(* Logix 5000 project; controller MV vendor 1 type 14 code 217 rev 31.11; software revision 31.00; part 40 of 53 *)
(* tags used below, declared in another part *)
   active : BOOL;
   MV_B100 : INT[255];   // AT FLAGS
   MV_N101 : INT[255];   // AT INT Fermentation control integer workspace
   MV_N110 : INT[255];   // MV DATA 0 CURRENT FV DATA
   MV_N12 : INT[255];   // SYS_PARMS System Parameter Fil e
   MV_N14 : INT[255];   // ME>PLC Inter PLC comms traf fic outbound
   MV_N7 : INT[255];   // INTEGER
   MV_SFile : INT[255];   // SLC Equivalent System File, So Original Code Can Remain
   MV_T102 : TIMER[10];
   MV_T4 : TIMER[20];
   MV_TENTH_HOUR_OUTPUT_BIT : BOOL;
   temp : INT;
(* MV_Common, continued *)

ROUTINE MV_FV_ELAPSED_102   (* ladder *)
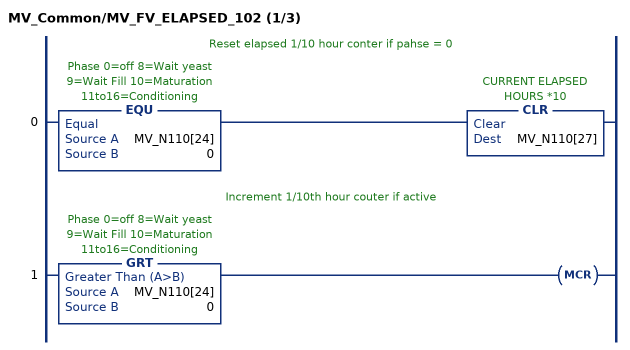
   // Reset elapsed 1/10 hour conter if pahse = 0
   0: EQU(MV_N110[24],0)CLR(MV_N110[27]);
   // Increment 1/10th hour couter if active
   1: GRT(MV_N110[24],0)MCR();
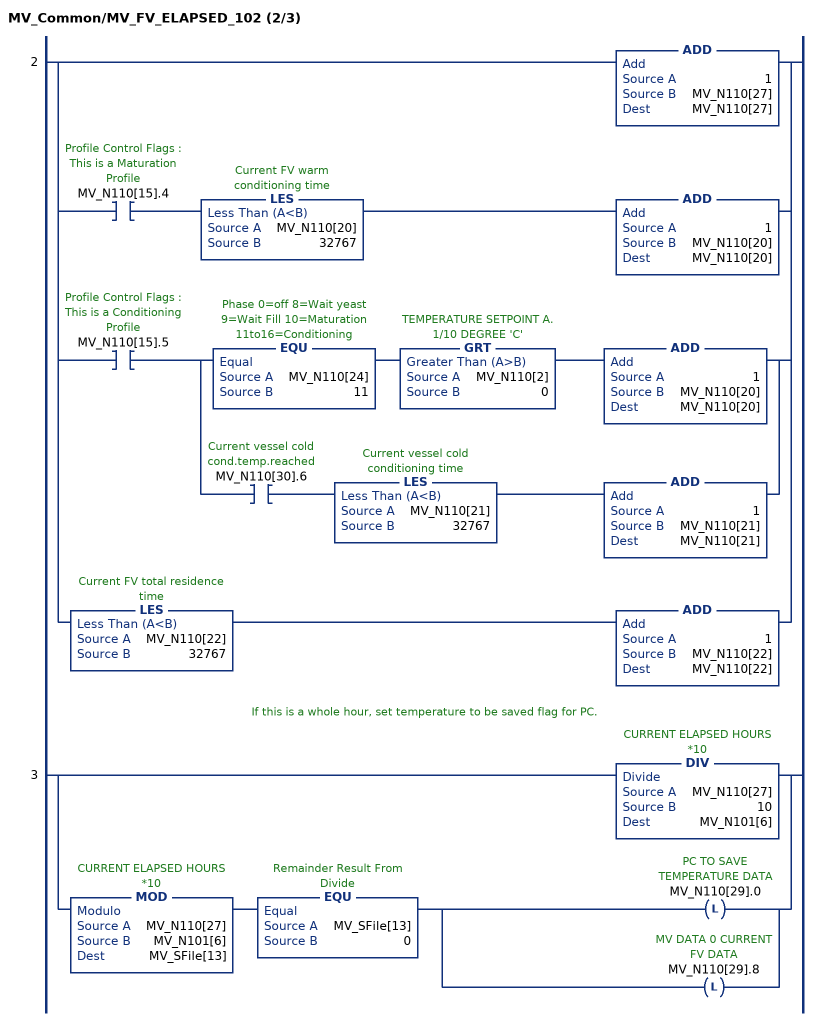
   2: [ADD(1,MV_N110[27],MV_N110[27]) ,XIC(MV_N110[15].4) LES(MV_N110[20],32767) ADD(1,MV_N110[20],MV_N110[20]) ,XIC(MV_N110[15].5) [EQU(MV_N110[24],11) GRT(MV_N110[2],0) ADD(1,MV_N110[20],MV_N110[20]) ,XIC(MV_N110[30].6) LES(MV_N110[21],32767) ADD(1,MV_N110[21],MV_N110[21]) ] ,LES(MV_N110[22],32767) ADD(1,MV_N110[22],MV_N110[22]) ];
   // If this is a whole hour, set temperature to be saved flag for PC.
   3: [DIV(MV_N110[27],10,MV_N101[6]) ,MOD(MV_N110[27],MV_N101[6],MV_SFile[13]) EQU(MV_SFile[13],0) [OTL(MV_N110[29].0) ,OTL(MV_N110[29].8) ] ];
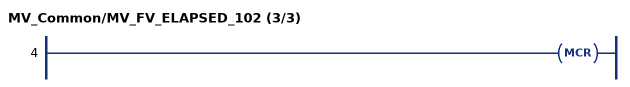
   4: MCR();
END_ROUTINE

ROUTINE MV_FV_MCP_100   (* ladder *)
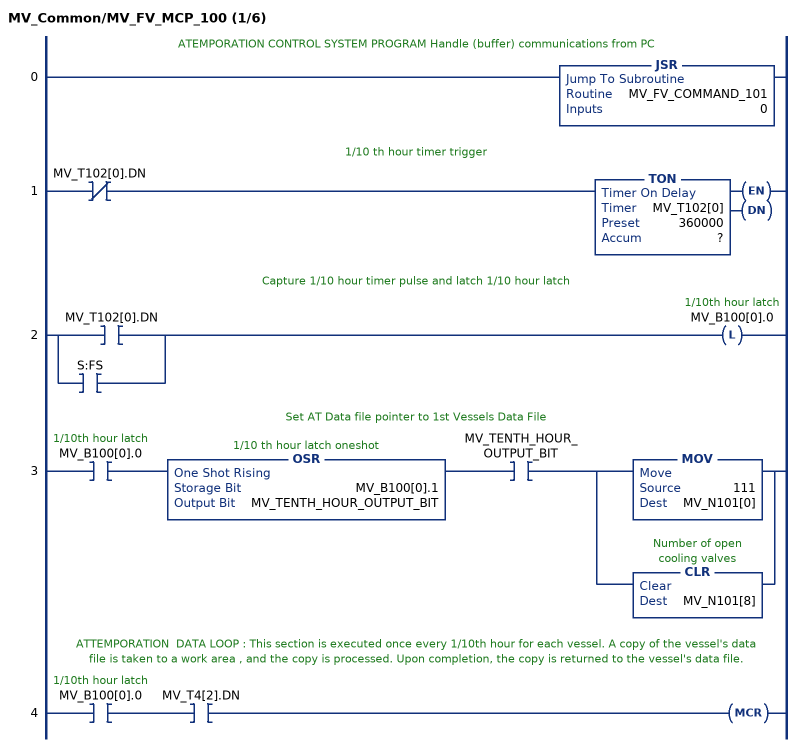
   // ATEMPORATION CONTROL SYSTEM PROGRAM Handle (buffer) communications from PC
   0: JSR(MV_FV_COMMAND_101,0);
   // 1/10 th hour timer trigger
   1: XIO(MV_T102[0].DN)TON(MV_T102[0],?,?);
   // Capture 1/10 hour timer pulse and latch 1/10 hour latch
   2: [XIC(MV_T102[0].DN) ,XIC(S:FS) ]OTL(MV_B100[0].0);
   // Set AT Data file pointer to 1st Vessels Data File
   3: XIC(MV_B100[0].0)OSR(MV_B100[0].1,MV_TENTH_HOUR_OUTPUT_BIT)XIC(MV_TENTH_HOUR_OUTPUT_BIT)[MOV(111,MV_N101[0]) ,CLR(MV_N101[8]) ];
   // ATTEMPORATION  DATA LOOP : This section is executed once every 1/10th hour for each vessel. A copy of the vessel's data file is taken to a work area , and the copy is processed. Upon completion, the copy is returned to the vessel's data file.
   4: XIC(MV_B100[0].0)XIC(MV_T4[2].DN)MCR();
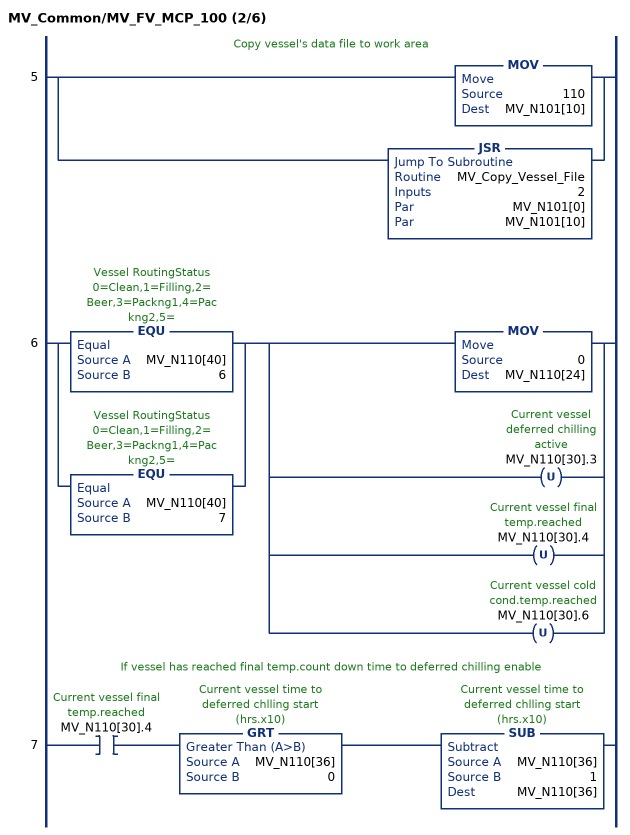
   // Copy vessel's data file to work area
   5: [MOV(110,MV_N101[10]) ,JSR(MV_Copy_Vessel_File,2,MV_N101[0],MV_N101[10]) ];
   6: [EQU(MV_N110[40],6) ,EQU(MV_N110[40],7) ][MOV(0,MV_N110[24]) ,OTU(MV_N110[30].3) ,OTU(MV_N110[30].4) ,OTU(MV_N110[30].6) ];
   // If vessel has reached final temp.count down time to deferred chilling enable
   7: XIC(MV_N110[30].4)GRT(MV_N110[36],0)SUB(MV_N110[36],1,MV_N110[36]);
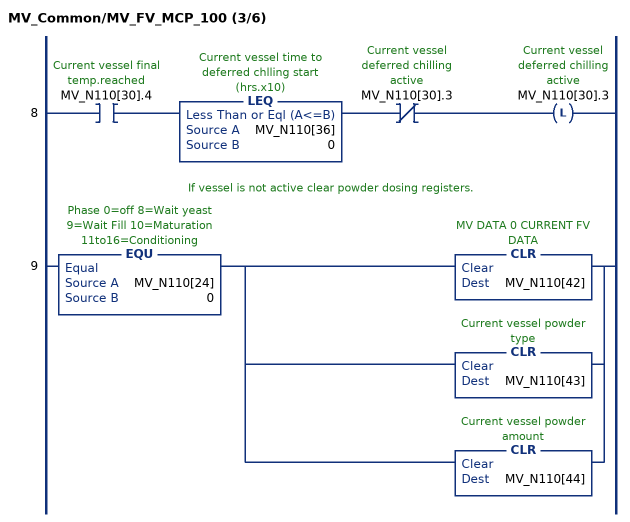
   8: XIC(MV_N110[30].4)LEQ(MV_N110[36],0)XIO(MV_N110[30].3)OTL(MV_N110[30].3);
   // If vessel is not active clear powder dosing registers.
   9: EQU(MV_N110[24],0)[CLR(MV_N110[42]) ,CLR(MV_N110[43]) ,CLR(MV_N110[44]) ];
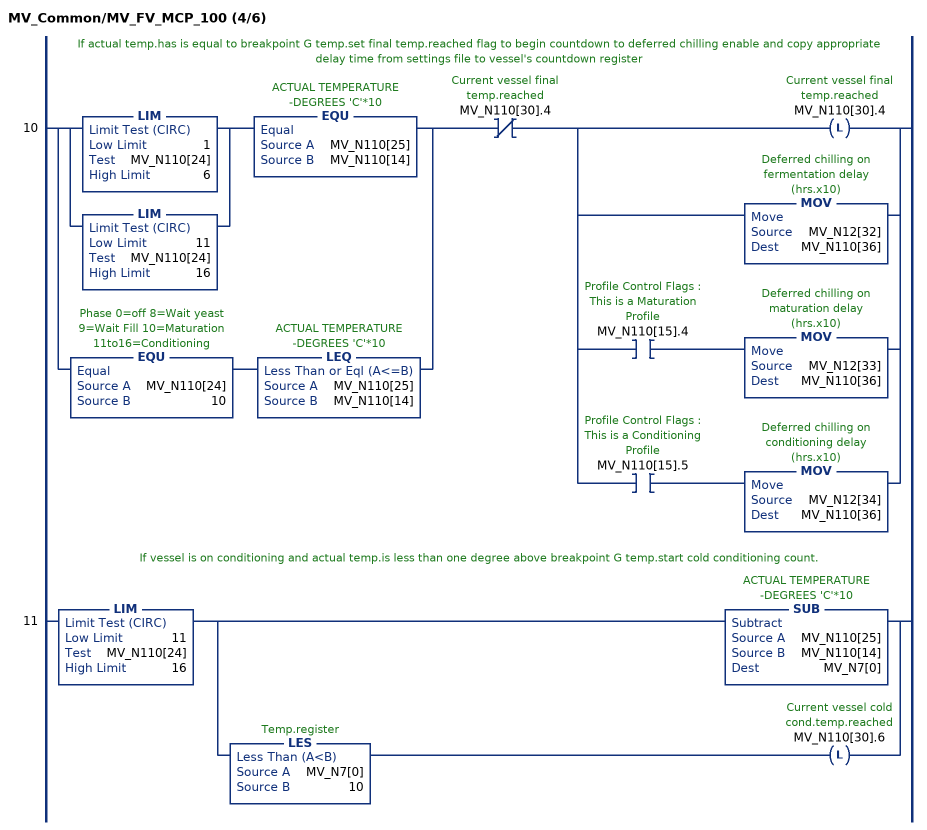
   // If actual temp.has is equal to breakpoint G temp.set final temp.reached flag to begin countdown to deferred chilling enable and copy appropriate delay time from settings file to vessel's countdown register
   10: [[LIM(1,MV_N110[24],6) ,LIM(11,MV_N110[24],16) ] EQU(MV_N110[25],MV_N110[14]) ,EQU(MV_N110[24],10) LEQ(MV_N110[25],MV_N110[14]) ]XIO(MV_N110[30].4)[OTL(MV_N110[30].4) ,MOV(MV_N12[32],MV_N110[36]) ,XIC(MV_N110[15].4) MOV(MV_N12[33],MV_N110[36]) ,XIC(MV_N110[15].5) MOV(MV_N12[34],MV_N110[36]) ];
   // If vessel is on conditioning and actual temp.is less than one degree above breakpoint G temp.start cold conditioning count.
   11: LIM(11,MV_N110[24],16)[SUB(MV_N110[25],MV_N110[14],MV_N7[0]) ,LES(MV_N7[0],10) OTL(MV_N110[30].6) ];
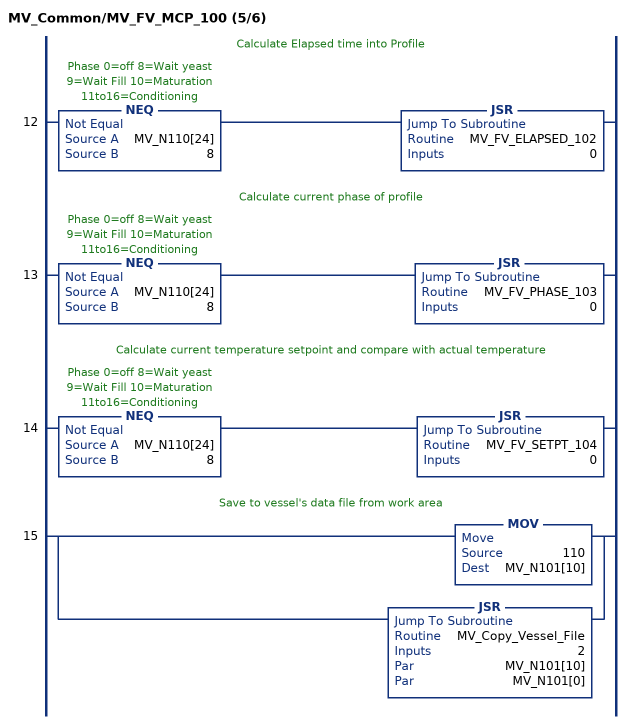
   // Calculate Elapsed time into Profile
   12: NEQ(MV_N110[24],8)JSR(MV_FV_ELAPSED_102,0);
   // Calculate current phase of profile
   13: NEQ(MV_N110[24],8)JSR(MV_FV_PHASE_103,0);
   // Calculate current temperature setpoint and compare with actual temperature
   14: NEQ(MV_N110[24],8)JSR(MV_FV_SETPT_104,0);
   // Save to vessel's data file from work area
   15: [MOV(110,MV_N101[10]) ,JSR(MV_Copy_Vessel_File,2,MV_N101[10],MV_N101[0]) ];
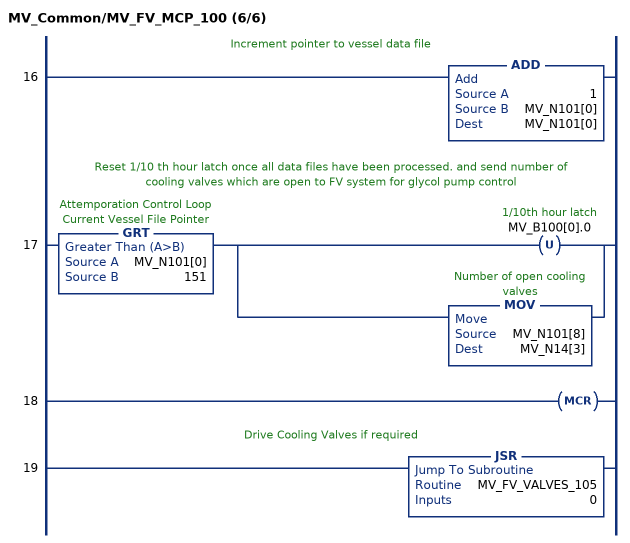
   // Increment pointer to vessel data file
   16: ADD(1,MV_N101[0],MV_N101[0]);
   // Reset 1/10 th hour latch once all data files have been processed. and send number of cooling valves which are open to FV system for glycol pump control
   17: GRT(MV_N101[0],151)[OTU(MV_B100[0].0) ,MOV(MV_N101[8],MV_N14[3]) ];
   18: MCR();
   // Drive Cooling Valves if required
   19: JSR(MV_FV_VALVES_105,0);
END_ROUTINE

ROUTINE MV_FV_PHASE_103   (* ladder *)
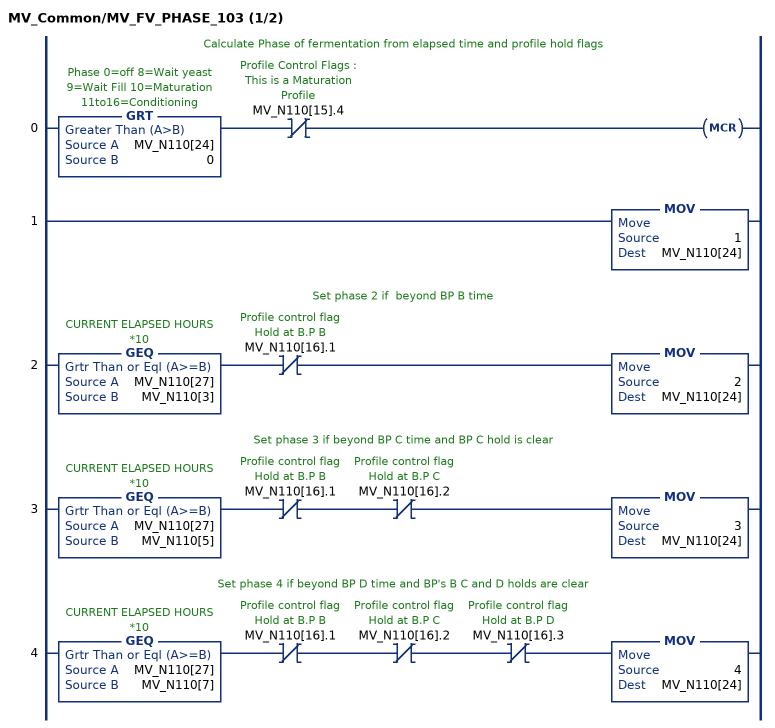
   // Calculate Phase of fermentation from elapsed time and profile hold flags
   0: GRT(MV_N110[24],0)XIO(MV_N110[15].4)MCR();
   1: MOV(1,MV_N110[24]);
   // Set phase 2 if  beyond BP B time
   2: GEQ(MV_N110[27],MV_N110[3])XIO(MV_N110[16].1)MOV(2,MV_N110[24]);
   // Set phase 3 if beyond BP C time and BP C hold is clear
   3: GEQ(MV_N110[27],MV_N110[5])XIO(MV_N110[16].1)XIO(MV_N110[16].2)MOV(3,MV_N110[24]);
   // Set phase 4 if beyond BP D time and BP's B C and D holds are clear
   4: GEQ(MV_N110[27],MV_N110[7])XIO(MV_N110[16].1)XIO(MV_N110[16].2)XIO(MV_N110[16].3)MOV(4,MV_N110[24]);
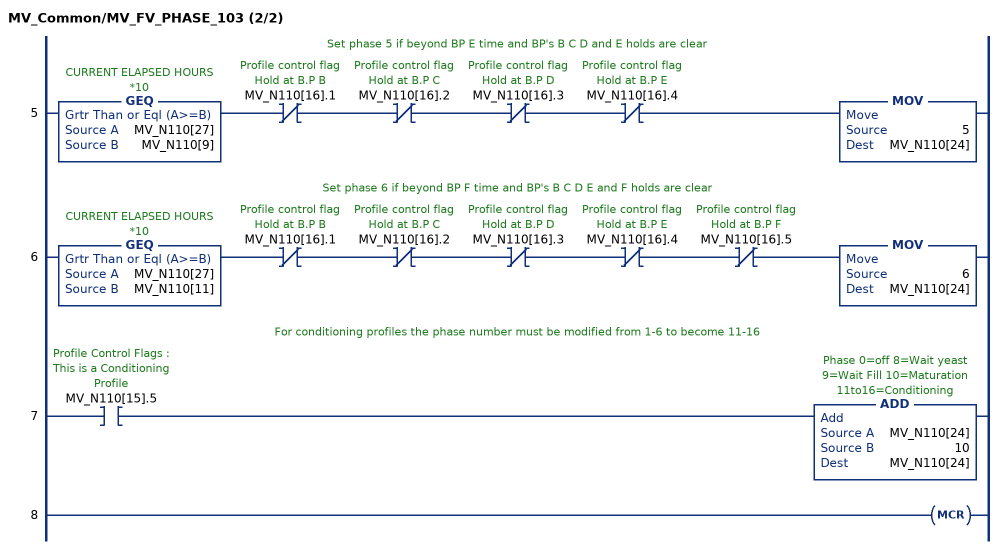
   // Set phase 5 if beyond BP E time and BP's B C D and E holds are clear
   5: GEQ(MV_N110[27],MV_N110[9])XIO(MV_N110[16].1)XIO(MV_N110[16].2)XIO(MV_N110[16].3)XIO(MV_N110[16].4)MOV(5,MV_N110[24]);
   // Set phase 6 if beyond BP F time and BP's B C D E and F holds are clear
   6: GEQ(MV_N110[27],MV_N110[11])XIO(MV_N110[16].1)XIO(MV_N110[16].2)XIO(MV_N110[16].3)XIO(MV_N110[16].4)XIO(MV_N110[16].5)MOV(6,MV_N110[24]);
   // For conditioning profiles the phase number must be modified from 1-6 to become 11-16
   7: XIC(MV_N110[15].5)ADD(MV_N110[24],10,MV_N110[24]);
   8: MCR();
END_ROUTINE

ROUTINE MV_FV_SETPT_104   (* ladder *)
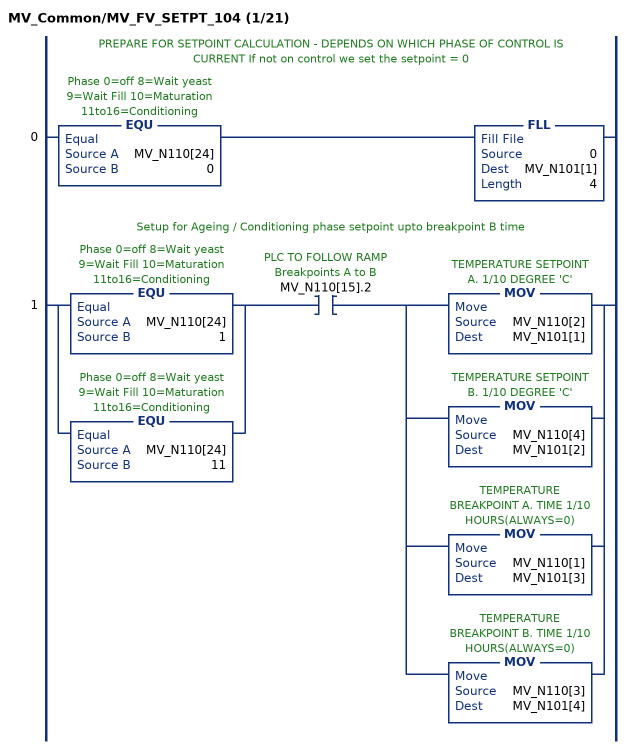
   // PREPARE FOR SETPOINT CALCULATION - DEPENDS ON WHICH PHASE OF CONTROL IS CURRENT If not on control we set the setpoint = 0
   0: EQU(MV_N110[24],0)FLL(0,MV_N101[1],4);
   // Setup for Ageing / Conditioning phase setpoint upto breakpoint B time
   1: [EQU(MV_N110[24],1) ,EQU(MV_N110[24],11) ]XIC(MV_N110[15].2)[MOV(MV_N110[2],MV_N101[1]) ,MOV(MV_N110[4],MV_N101[2]) ,MOV(MV_N110[1],MV_N101[3]) ,MOV(MV_N110[3],MV_N101[4]) ];
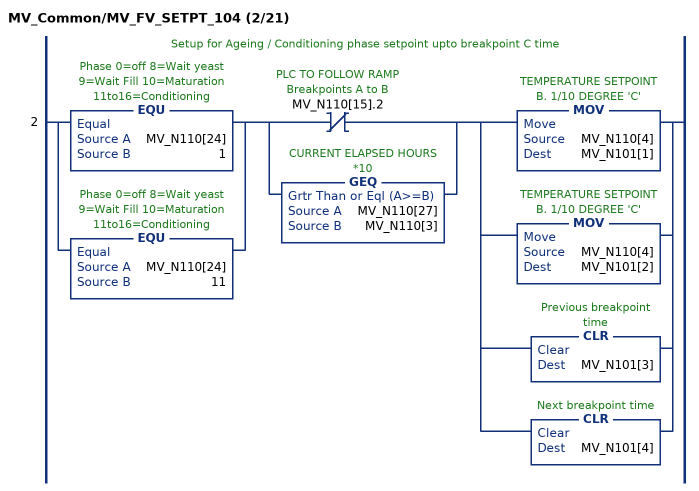
   // Setup for Ageing / Conditioning phase setpoint upto breakpoint C time
   2: [EQU(MV_N110[24],1) ,EQU(MV_N110[24],11) ][XIO(MV_N110[15].2) ,GEQ(MV_N110[27],MV_N110[3]) ][MOV(MV_N110[4],MV_N101[1]) ,MOV(MV_N110[4],MV_N101[2]) ,CLR(MV_N101[3]) ,CLR(MV_N101[4]) ];
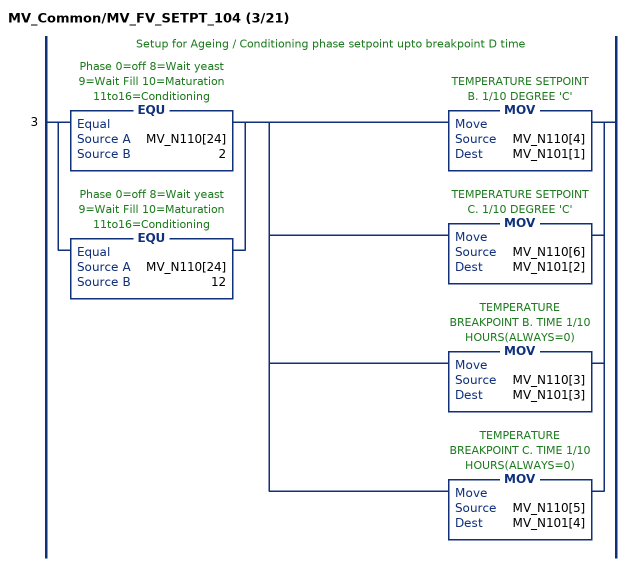
   // Setup for Ageing / Conditioning phase setpoint upto breakpoint D time
   3: [EQU(MV_N110[24],2) ,EQU(MV_N110[24],12) ][MOV(MV_N110[4],MV_N101[1]) ,MOV(MV_N110[6],MV_N101[2]) ,MOV(MV_N110[3],MV_N101[3]) ,MOV(MV_N110[5],MV_N101[4]) ];
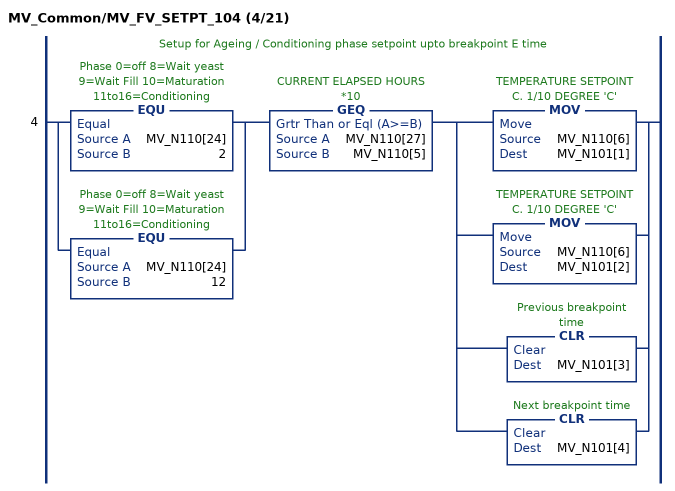
   // Setup for Ageing / Conditioning phase setpoint upto breakpoint E time
   4: [EQU(MV_N110[24],2) ,EQU(MV_N110[24],12) ]GEQ(MV_N110[27],MV_N110[5])[MOV(MV_N110[6],MV_N101[1]) ,MOV(MV_N110[6],MV_N101[2]) ,CLR(MV_N101[3]) ,CLR(MV_N101[4]) ];
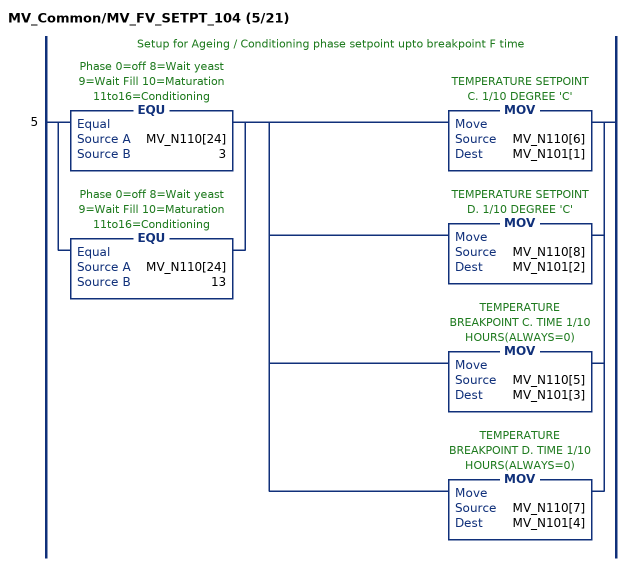
   // Setup for Ageing / Conditioning phase setpoint upto breakpoint F time
   5: [EQU(MV_N110[24],3) ,EQU(MV_N110[24],13) ][MOV(MV_N110[6],MV_N101[1]) ,MOV(MV_N110[8],MV_N101[2]) ,MOV(MV_N110[5],MV_N101[3]) ,MOV(MV_N110[7],MV_N101[4]) ];
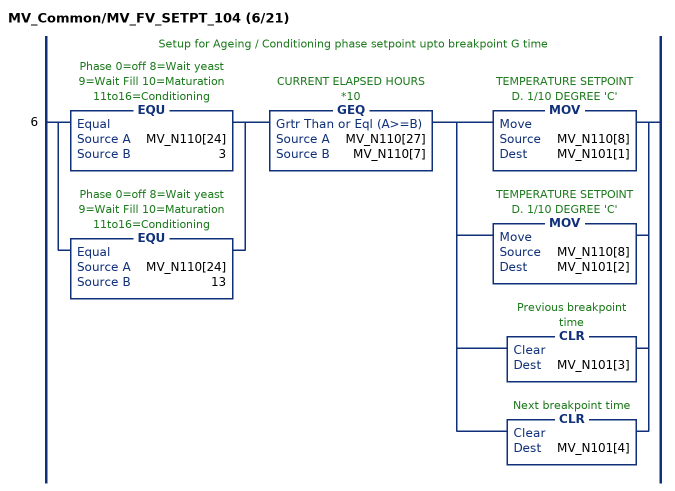
   // Setup for Ageing / Conditioning phase setpoint upto breakpoint G time
   6: [EQU(MV_N110[24],3) ,EQU(MV_N110[24],13) ]GEQ(MV_N110[27],MV_N110[7])[MOV(MV_N110[8],MV_N101[1]) ,MOV(MV_N110[8],MV_N101[2]) ,CLR(MV_N101[3]) ,CLR(MV_N101[4]) ];
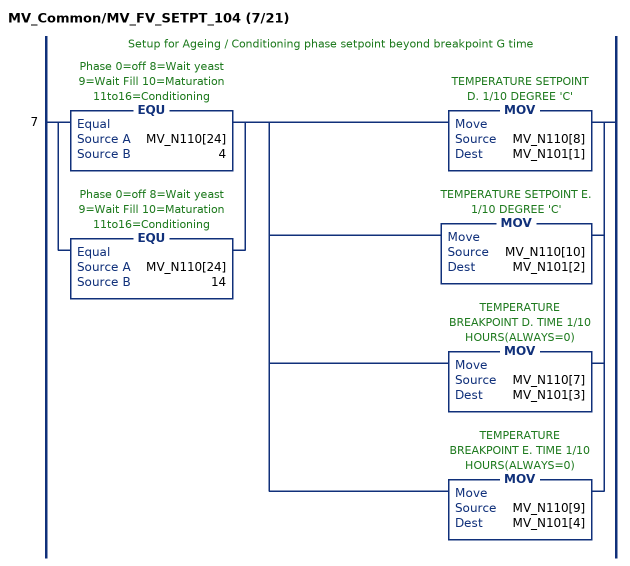
   // Setup for Ageing / Conditioning phase setpoint beyond breakpoint G time
   7: [EQU(MV_N110[24],4) ,EQU(MV_N110[24],14) ][MOV(MV_N110[8],MV_N101[1]) ,MOV(MV_N110[10],MV_N101[2]) ,MOV(MV_N110[7],MV_N101[3]) ,MOV(MV_N110[9],MV_N101[4]) ];
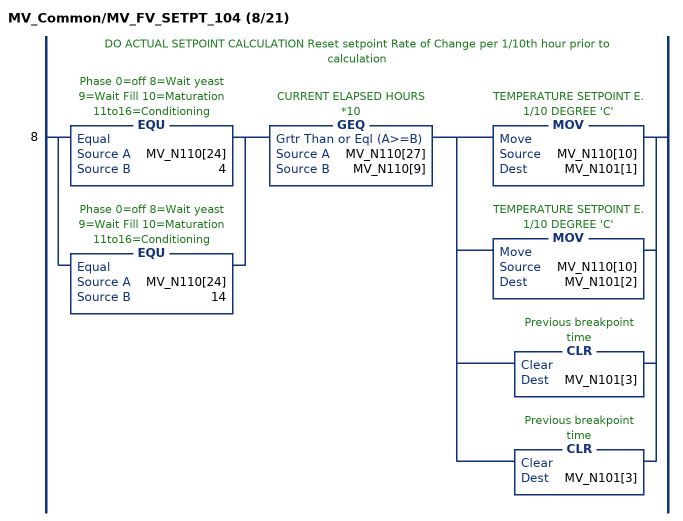
   // DO ACTUAL SETPOINT CALCULATION Reset setpoint Rate of Change per 1/10th hour prior to calculation
   8: [EQU(MV_N110[24],4) ,EQU(MV_N110[24],14) ]GEQ(MV_N110[27],MV_N110[9])[MOV(MV_N110[10],MV_N101[1]) ,MOV(MV_N110[10],MV_N101[2]) ,CLR(MV_N101[3]) ,CLR(MV_N101[3]) ];
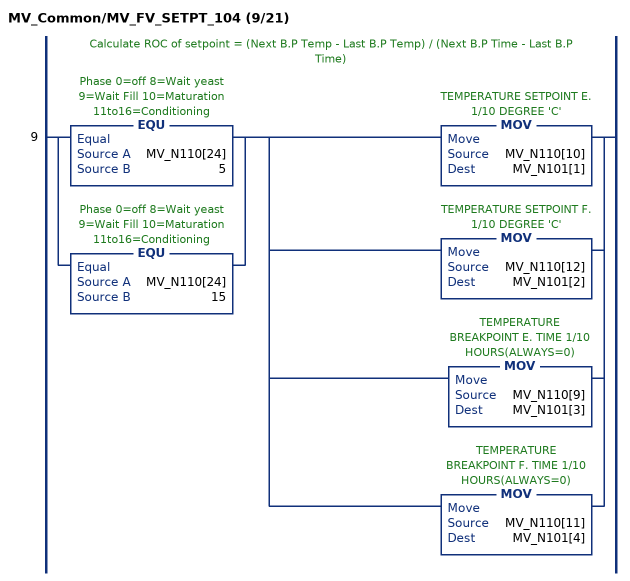
   // Calculate ROC of setpoint = (Next B.P Temp - Last B.P Temp) / (Next B.P Time - Last B.P Time)
   9: [EQU(MV_N110[24],5) ,EQU(MV_N110[24],15) ][MOV(MV_N110[10],MV_N101[1]) ,MOV(MV_N110[12],MV_N101[2]) ,MOV(MV_N110[9],MV_N101[3]) ,MOV(MV_N110[11],MV_N101[4]) ];
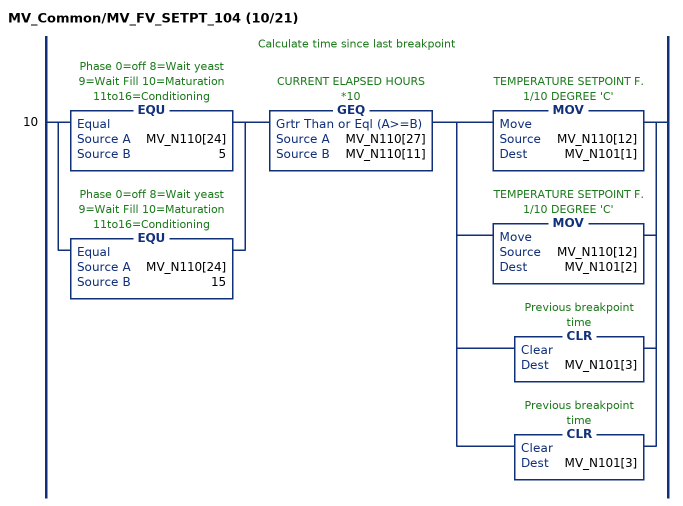
   // Calculate time since last breakpoint
   10: [EQU(MV_N110[24],5) ,EQU(MV_N110[24],15) ]GEQ(MV_N110[27],MV_N110[11])[MOV(MV_N110[12],MV_N101[1]) ,MOV(MV_N110[12],MV_N101[2]) ,CLR(MV_N101[3]) ,CLR(MV_N101[3]) ];
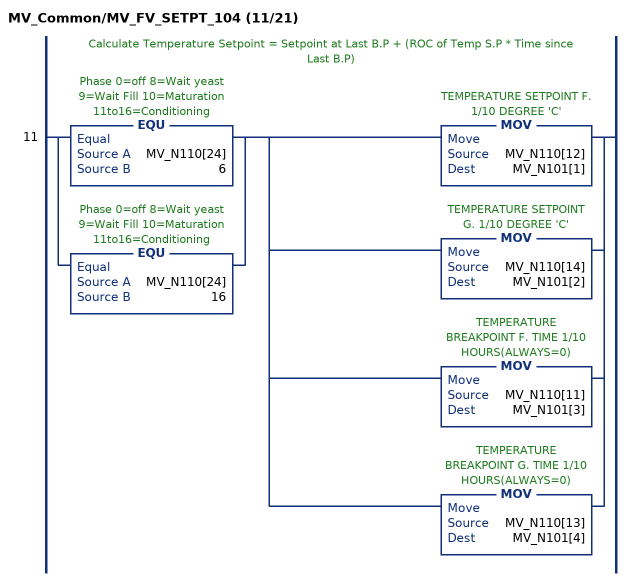
   // Calculate Temperature Setpoint = Setpoint at Last B.P + (ROC of Temp S.P * Time since Last B.P)
   11: [EQU(MV_N110[24],6) ,EQU(MV_N110[24],16) ][MOV(MV_N110[12],MV_N101[1]) ,MOV(MV_N110[14],MV_N101[2]) ,MOV(MV_N110[11],MV_N101[3]) ,MOV(MV_N110[13],MV_N101[4]) ];
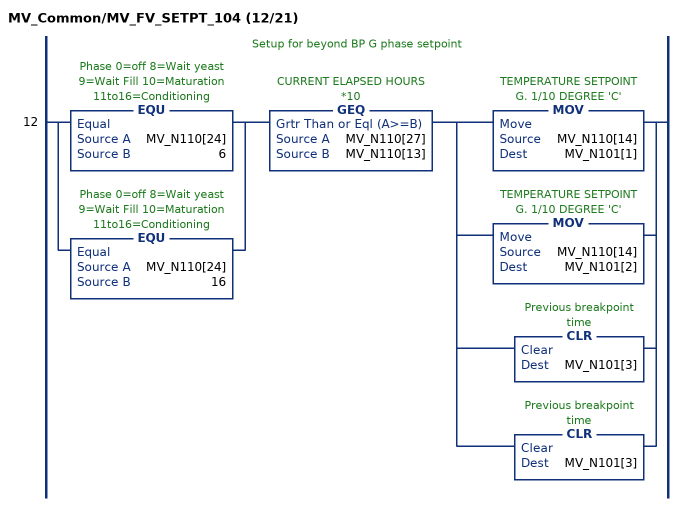
   // Setup for beyond BP G phase setpoint
   12: [EQU(MV_N110[24],6) ,EQU(MV_N110[24],16) ]GEQ(MV_N110[27],MV_N110[13])[MOV(MV_N110[14],MV_N101[1]) ,MOV(MV_N110[14],MV_N101[2]) ,CLR(MV_N101[3]) ,CLR(MV_N101[3]) ];
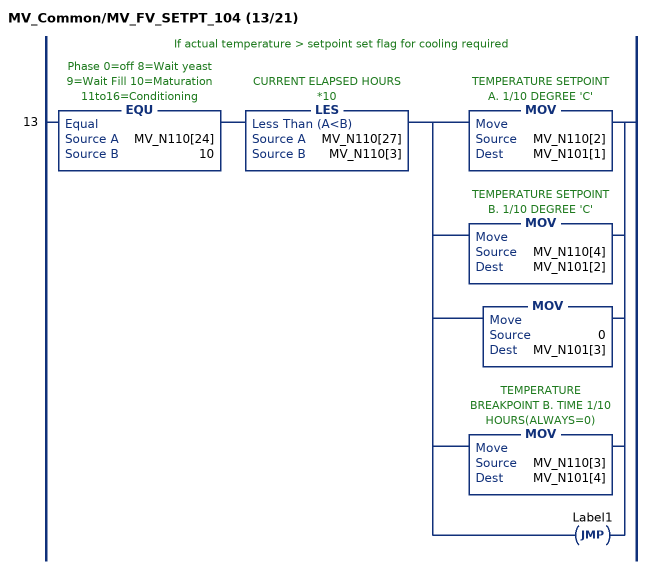
   // If actual temperature > setpoint set flag for cooling required
   13: EQU(MV_N110[24],10)LES(MV_N110[27],MV_N110[3])[MOV(MV_N110[2],MV_N101[1]) ,MOV(MV_N110[4],MV_N101[2]) ,MOV(0,MV_N101[3]) ,MOV(MV_N110[3],MV_N101[4]) ,JMP(Label1) ];
